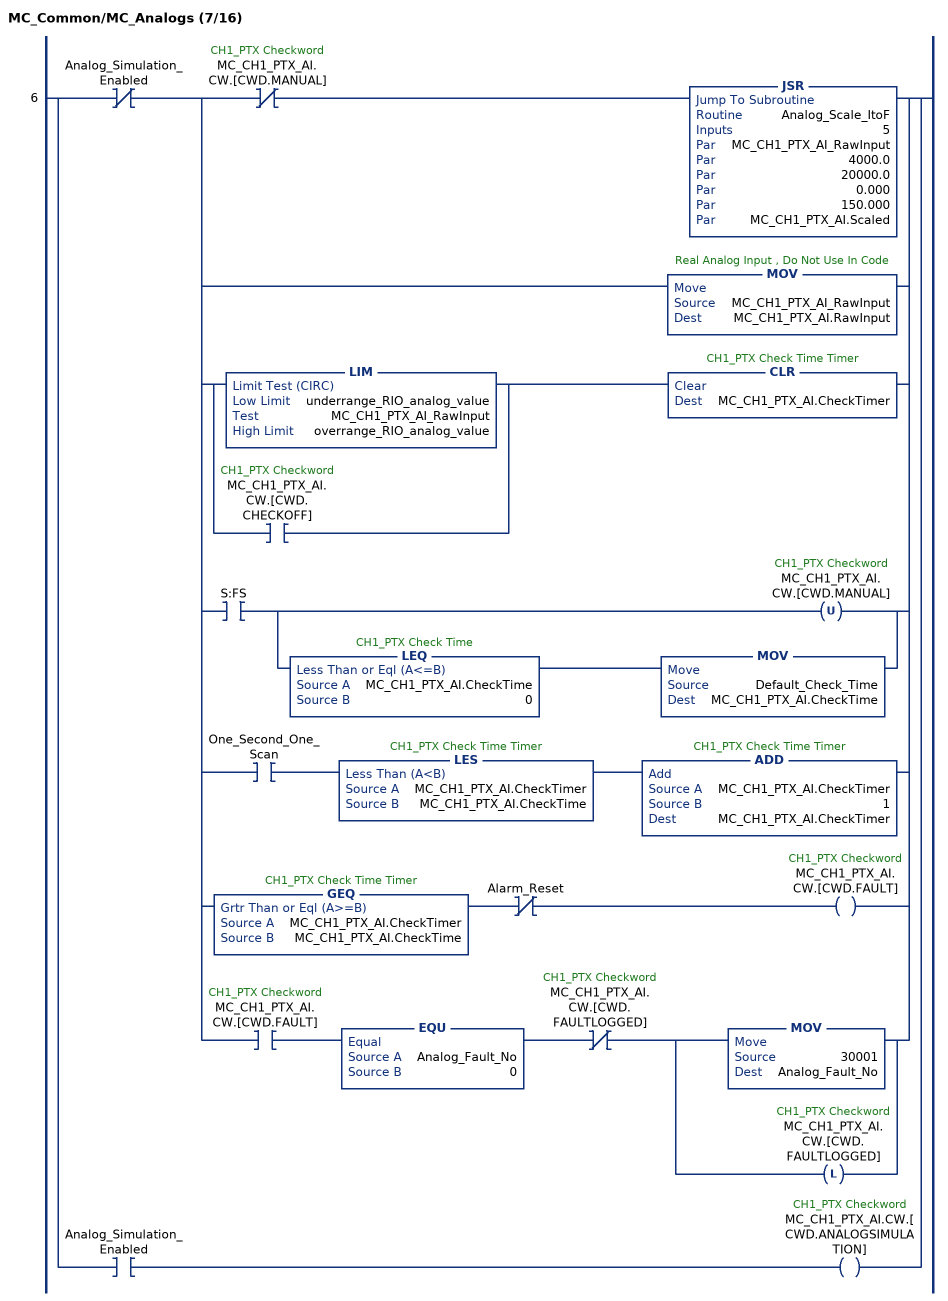
   6: [XIO(Analog_Simulation_Enabled) [XIO(MC_CH1_PTX_AI.CW.[CWD.MANUAL]) JSR(Analog_Scale_ItoF,5,MC_CH1_PTX_AI_RawInput,4000.0,20000.0,0.000,150.000,MC_CH1_PTX_AI.Scaled) ,MOV(MC_CH1_PTX_AI_RawInput,MC_CH1_PTX_AI.RawInput) ,[LIM(underrange_RIO_analog_value,MC_CH1_PTX_AI_RawInput,overrange_RIO_analog_value) ,XIC(MC_CH1_PTX_AI.CW.[CWD.CHECKOFF]) ] CLR(MC_CH1_PTX_AI.CheckTimer) ,XIC(S:FS) [OTU(MC_CH1_PTX_AI.CW.[CWD.MANUAL]) ,LEQ(MC_CH1_PTX_AI.CheckTime,0) MOV(Default_Check_Time,MC_CH1_PTX_AI.CheckTime) ] ,XIC(One_Second_One_Scan) LES(MC_CH1_PTX_AI.CheckTimer,MC_CH1_PTX_AI.CheckTime) ADD(MC_CH1_PTX_AI.CheckTimer,1,MC_CH1_PTX_AI.CheckTimer) ,GEQ(MC_CH1_PTX_AI.CheckTimer,MC_CH1_PTX_AI.CheckTime) XIO(Alarm_Reset) OTE(MC_CH1_PTX_AI.CW.[CWD.FAULT]) ,XIC(MC_CH1_PTX_AI.CW.[CWD.FAULT]) EQU(Analog_Fault_No,0) XIO(MC_CH1_PTX_AI.CW.[CWD.FAULTLOGGED]) [MOV(30001,Analog_Fault_No) ,OTL(MC_CH1_PTX_AI.CW.[CWD.FAULTLOGGED]) ] ] ,XIC(Analog_Simulation_Enabled) OTE(MC_CH1_PTX_AI.CW.[CWD.ANALOGSIMULATION]) ];
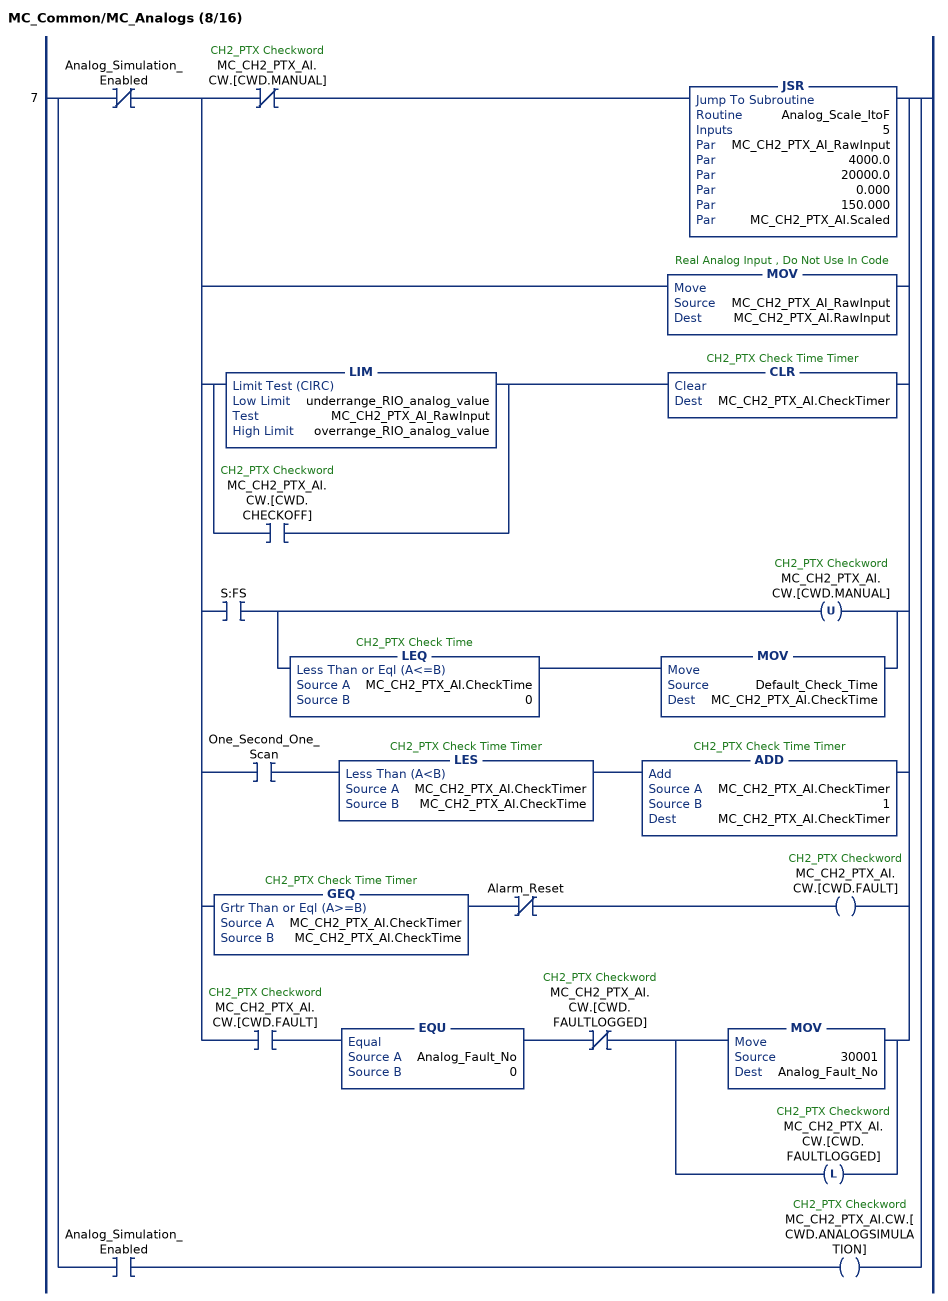
   7: [XIO(Analog_Simulation_Enabled) [XIO(MC_CH2_PTX_AI.CW.[CWD.MANUAL]) JSR(Analog_Scale_ItoF,5,MC_CH2_PTX_AI_RawInput,4000.0,20000.0,0.000,150.000,MC_CH2_PTX_AI.Scaled) ,MOV(MC_CH2_PTX_AI_RawInput,MC_CH2_PTX_AI.RawInput) ,[LIM(underrange_RIO_analog_value,MC_CH2_PTX_AI_RawInput,overrange_RIO_analog_value) ,XIC(MC_CH2_PTX_AI.CW.[CWD.CHECKOFF]) ] CLR(MC_CH2_PTX_AI.CheckTimer) ,XIC(S:FS) [OTU(MC_CH2_PTX_AI.CW.[CWD.MANUAL]) ,LEQ(MC_CH2_PTX_AI.CheckTime,0) MOV(Default_Check_Time,MC_CH2_PTX_AI.CheckTime) ] ,XIC(One_Second_One_Scan) LES(MC_CH2_PTX_AI.CheckTimer,MC_CH2_PTX_AI.CheckTime) ADD(MC_CH2_PTX_AI.CheckTimer,1,MC_CH2_PTX_AI.CheckTimer) ,GEQ(MC_CH2_PTX_AI.CheckTimer,MC_CH2_PTX_AI.CheckTime) XIO(Alarm_Reset) OTE(MC_CH2_PTX_AI.CW.[CWD.FAULT]) ,XIC(MC_CH2_PTX_AI.CW.[CWD.FAULT]) EQU(Analog_Fault_No,0) XIO(MC_CH2_PTX_AI.CW.[CWD.FAULTLOGGED]) [MOV(30001,Analog_Fault_No) ,OTL(MC_CH2_PTX_AI.CW.[CWD.FAULTLOGGED]) ] ] ,XIC(Analog_Simulation_Enabled) OTE(MC_CH2_PTX_AI.CW.[CWD.ANALOGSIMULATION]) ];
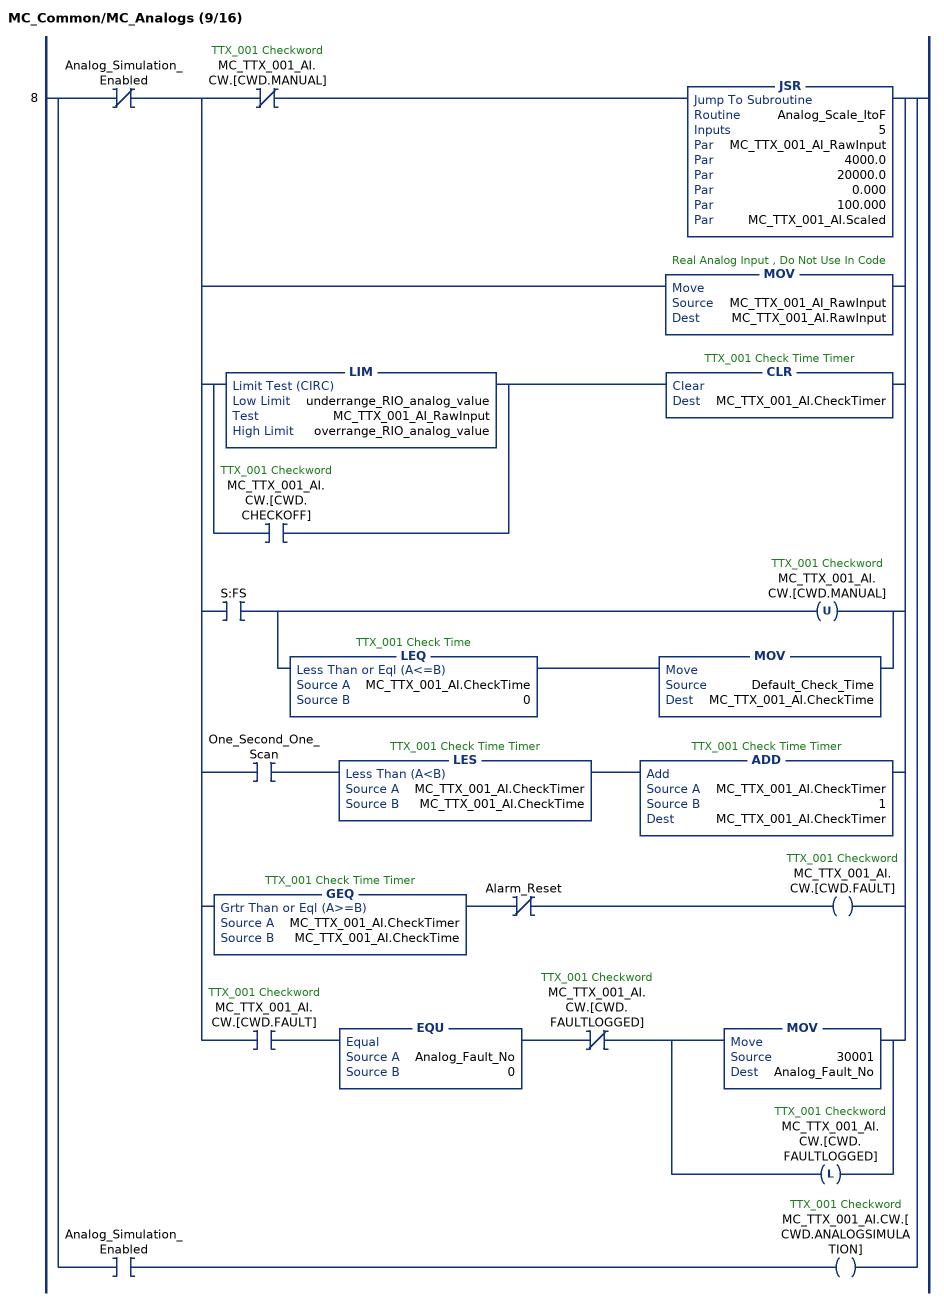
   8: [XIO(Analog_Simulation_Enabled) [XIO(MC_TTX_001_AI.CW.[CWD.MANUAL]) JSR(Analog_Scale_ItoF,5,MC_TTX_001_AI_RawInput,4000.0,20000.0,0.000,100.000,MC_TTX_001_AI.Scaled) ,MOV(MC_TTX_001_AI_RawInput,MC_TTX_001_AI.RawInput) ,[LIM(underrange_RIO_analog_value,MC_TTX_001_AI_RawInput,overrange_RIO_analog_value) ,XIC(MC_TTX_001_AI.CW.[CWD.CHECKOFF]) ] CLR(MC_TTX_001_AI.CheckTimer) ,XIC(S:FS) [OTU(MC_TTX_001_AI.CW.[CWD.MANUAL]) ,LEQ(MC_TTX_001_AI.CheckTime,0) MOV(Default_Check_Time,MC_TTX_001_AI.CheckTime) ] ,XIC(One_Second_One_Scan) LES(MC_TTX_001_AI.CheckTimer,MC_TTX_001_AI.CheckTime) ADD(MC_TTX_001_AI.CheckTimer,1,MC_TTX_001_AI.CheckTimer) ,GEQ(MC_TTX_001_AI.CheckTimer,MC_TTX_001_AI.CheckTime) XIO(Alarm_Reset) OTE(MC_TTX_001_AI.CW.[CWD.FAULT]) ,XIC(MC_TTX_001_AI.CW.[CWD.FAULT]) EQU(Analog_Fault_No,0) XIO(MC_TTX_001_AI.CW.[CWD.FAULTLOGGED]) [MOV(30001,Analog_Fault_No) ,OTL(MC_TTX_001_AI.CW.[CWD.FAULTLOGGED]) ] ] ,XIC(Analog_Simulation_Enabled) OTE(MC_TTX_001_AI.CW.[CWD.ANALOGSIMULATION]) ];
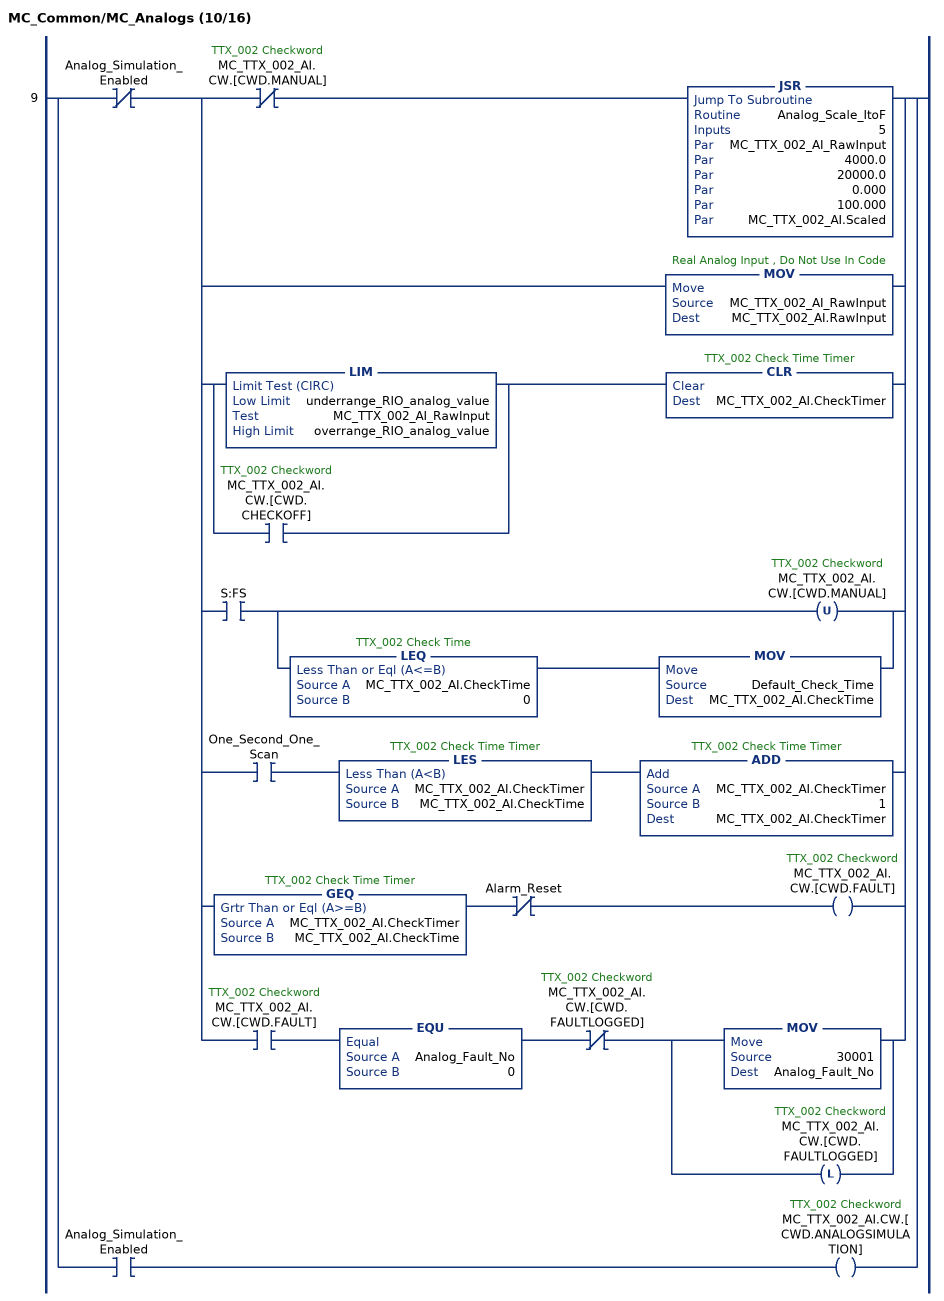
   9: [XIO(Analog_Simulation_Enabled) [XIO(MC_TTX_002_AI.CW.[CWD.MANUAL]) JSR(Analog_Scale_ItoF,5,MC_TTX_002_AI_RawInput,4000.0,20000.0,0.000,100.000,MC_TTX_002_AI.Scaled) ,MOV(MC_TTX_002_AI_RawInput,MC_TTX_002_AI.RawInput) ,[LIM(underrange_RIO_analog_value,MC_TTX_002_AI_RawInput,overrange_RIO_analog_value) ,XIC(MC_TTX_002_AI.CW.[CWD.CHECKOFF]) ] CLR(MC_TTX_002_AI.CheckTimer) ,XIC(S:FS) [OTU(MC_TTX_002_AI.CW.[CWD.MANUAL]) ,LEQ(MC_TTX_002_AI.CheckTime,0) MOV(Default_Check_Time,MC_TTX_002_AI.CheckTime) ] ,XIC(One_Second_One_Scan) LES(MC_TTX_002_AI.CheckTimer,MC_TTX_002_AI.CheckTime) ADD(MC_TTX_002_AI.CheckTimer,1,MC_TTX_002_AI.CheckTimer) ,GEQ(MC_TTX_002_AI.CheckTimer,MC_TTX_002_AI.CheckTime) XIO(Alarm_Reset) OTE(MC_TTX_002_AI.CW.[CWD.FAULT]) ,XIC(MC_TTX_002_AI.CW.[CWD.FAULT]) EQU(Analog_Fault_No,0) XIO(MC_TTX_002_AI.CW.[CWD.FAULTLOGGED]) [MOV(30001,Analog_Fault_No) ,OTL(MC_TTX_002_AI.CW.[CWD.FAULTLOGGED]) ] ] ,XIC(Analog_Simulation_Enabled) OTE(MC_TTX_002_AI.CW.[CWD.ANALOGSIMULATION]) ];
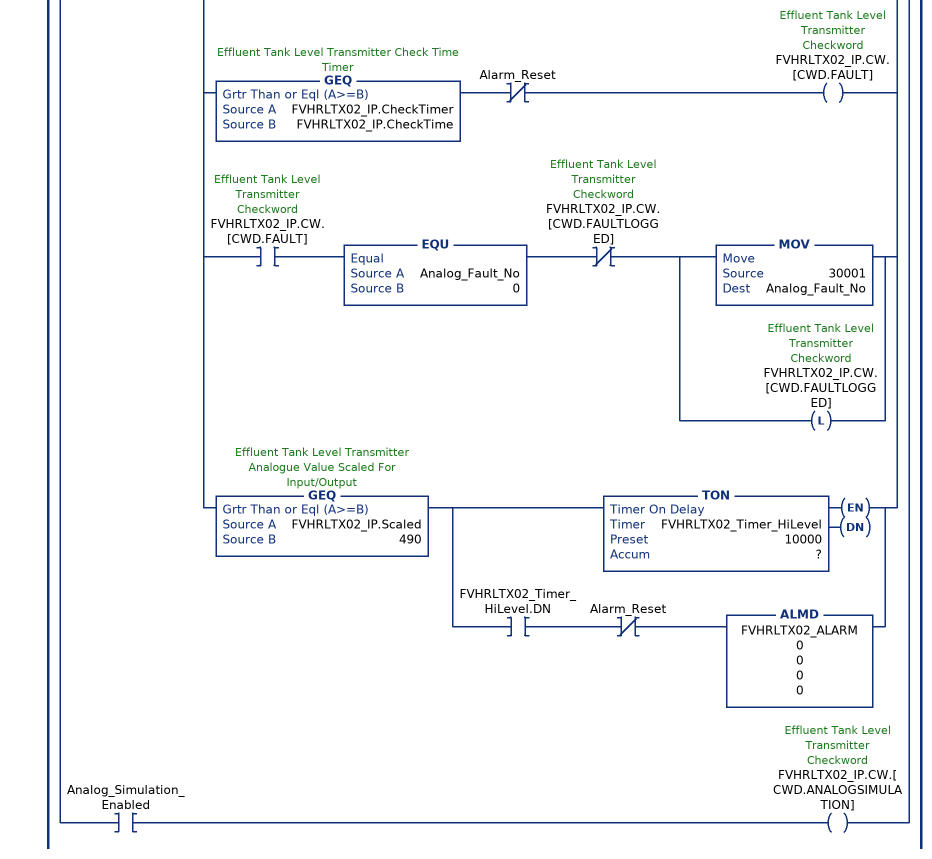
   10: [XIO(Analog_Simulation_Enabled) [XIO(FVHRLTX02_IP.CW.[CWD.MANUAL]) [JSR(Analog_Scale_ItoF,5,FVHRLTX02_IP_RawInput,4000.0,20000.0,0.0,500.0,FVHRLTX02_IP.Scaled) ,CPT(FVHRLTX02_IP_Percentage,(FVHRLTX02_IP.Scaled / 500) * 100) ] ,MOV(FVHRLTX02_IP_RawInput,FVHRLTX02_IP.RawInput) ,[LIM(underrange_RIO_analog_value,FVHRLTX02_IP_RawInput,overrange_RIO_analog_value) ,XIC(FVHRLTX02_IP.CW.[CWD.CHECKOFF]) ] CLR(FVHRLTX02_IP.CheckTimer) ,XIC(S:FS) [OTU(FVHRLTX02_IP.CW.[CWD.MANUAL]) ,LEQ(FVHRLTX02_IP.CheckTime,0) MOV(Default_Check_Time,FVHRLTX02_IP.CheckTime) ] ,XIC(One_Second_One_Scan) LES(FVHRLTX02_IP.CheckTimer,FVHRLTX02_IP.CheckTime) ADD(FVHRLTX02_IP.CheckTimer,1,FVHRLTX02_IP.CheckTimer) ,GEQ(FVHRLTX02_IP.CheckTimer,FVHRLTX02_IP.CheckTime) XIO(Alarm_Reset) OTE(FVHRLTX02_IP.CW.[CWD.FAULT]) ,XIC(FVHRLTX02_IP.CW.[CWD.FAULT]) EQU(Analog_Fault_No,0) XIO(FVHRLTX02_IP.CW.[CWD.FAULTLOGGED]) [MOV(30001,Analog_Fault_No) ,OTL(FVHRLTX02_IP.CW.[CWD.FAULTLOGGED]) ] ,GEQ(FVHRLTX02_IP.Scaled,490) [TON(FVHRLTX02_Timer_HiLevel,?,?) ,XIC(FVHRLTX02_Timer_HiLevel.DN) XIO(Alarm_Reset) ALMD(FVHRLTX02_ALARM,0,0,0,0) ] ] ,XIC(Analog_Simulation_Enabled) OTE(FVHRLTX02_IP.CW.[CWD.ANALOGSIMULATION]) ];
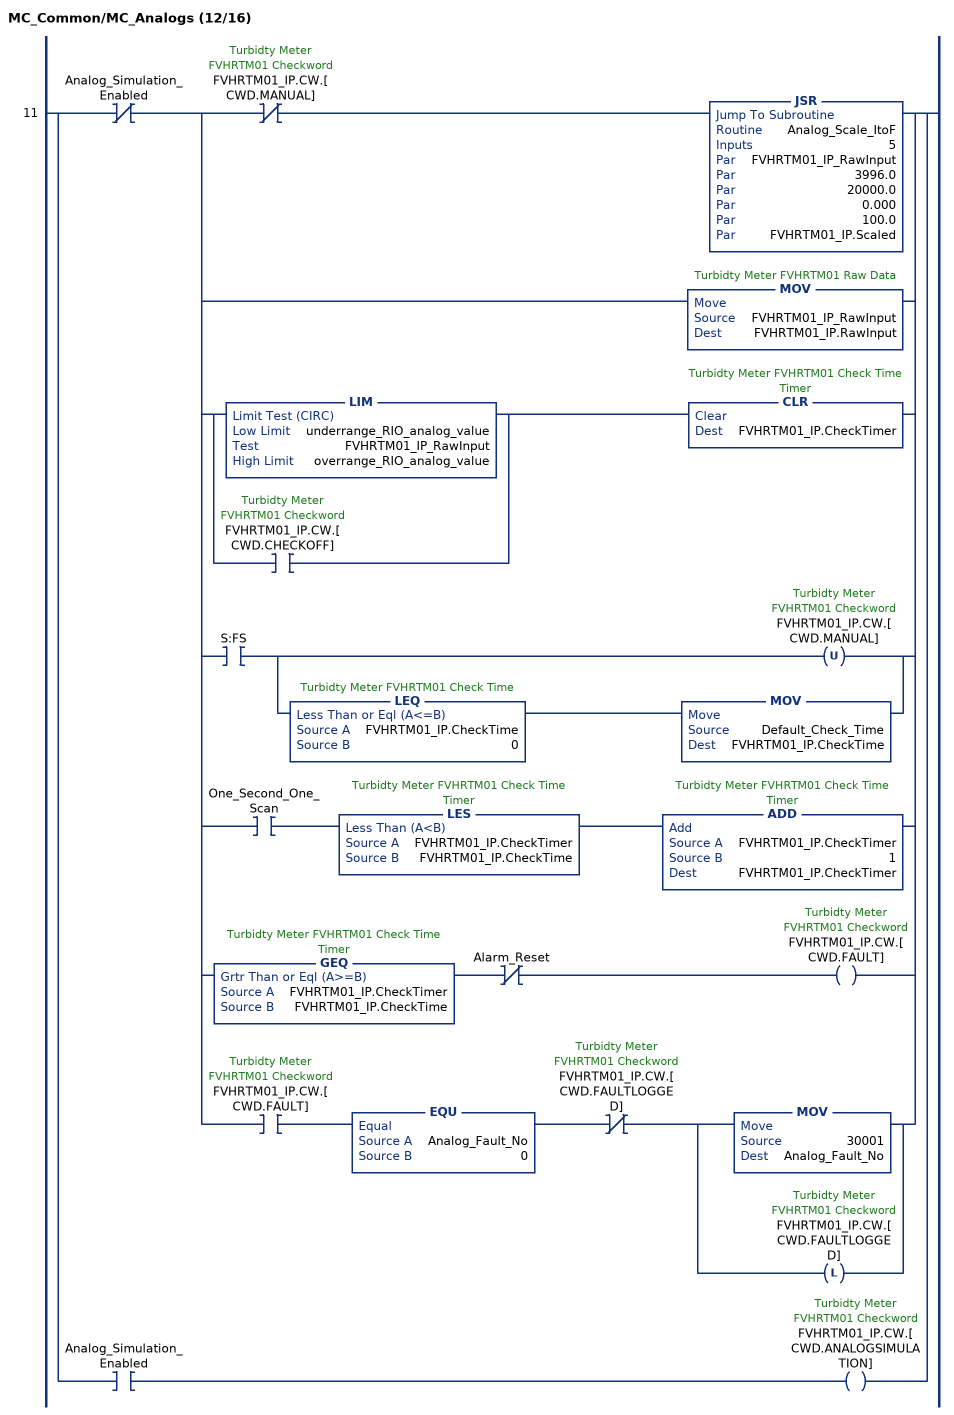
   11: [XIO(Analog_Simulation_Enabled) [XIO(FVHRTM01_IP.CW.[CWD.MANUAL]) JSR(Analog_Scale_ItoF,5,FVHRTM01_IP_RawInput,3996.0,20000.0,0.000,100.0,FVHRTM01_IP.Scaled) ,MOV(FVHRTM01_IP_RawInput,FVHRTM01_IP.RawInput) ,[LIM(underrange_RIO_analog_value,FVHRTM01_IP_RawInput,overrange_RIO_analog_value) ,XIC(FVHRTM01_IP.CW.[CWD.CHECKOFF]) ] CLR(FVHRTM01_IP.CheckTimer) ,XIC(S:FS) [OTU(FVHRTM01_IP.CW.[CWD.MANUAL]) ,LEQ(FVHRTM01_IP.CheckTime,0) MOV(Default_Check_Time,FVHRTM01_IP.CheckTime) ] ,XIC(One_Second_One_Scan) LES(FVHRTM01_IP.CheckTimer,FVHRTM01_IP.CheckTime) ADD(FVHRTM01_IP.CheckTimer,1,FVHRTM01_IP.CheckTimer) ,GEQ(FVHRTM01_IP.CheckTimer,FVHRTM01_IP.CheckTime) XIO(Alarm_Reset) OTE(FVHRTM01_IP.CW.[CWD.FAULT]) ,XIC(FVHRTM01_IP.CW.[CWD.FAULT]) EQU(Analog_Fault_No,0) XIO(FVHRTM01_IP.CW.[CWD.FAULTLOGGED]) [MOV(30001,Analog_Fault_No) ,OTL(FVHRTM01_IP.CW.[CWD.FAULTLOGGED]) ] ] ,XIC(Analog_Simulation_Enabled) OTE(FVHRTM01_IP.CW.[CWD.ANALOGSIMULATION]) ];
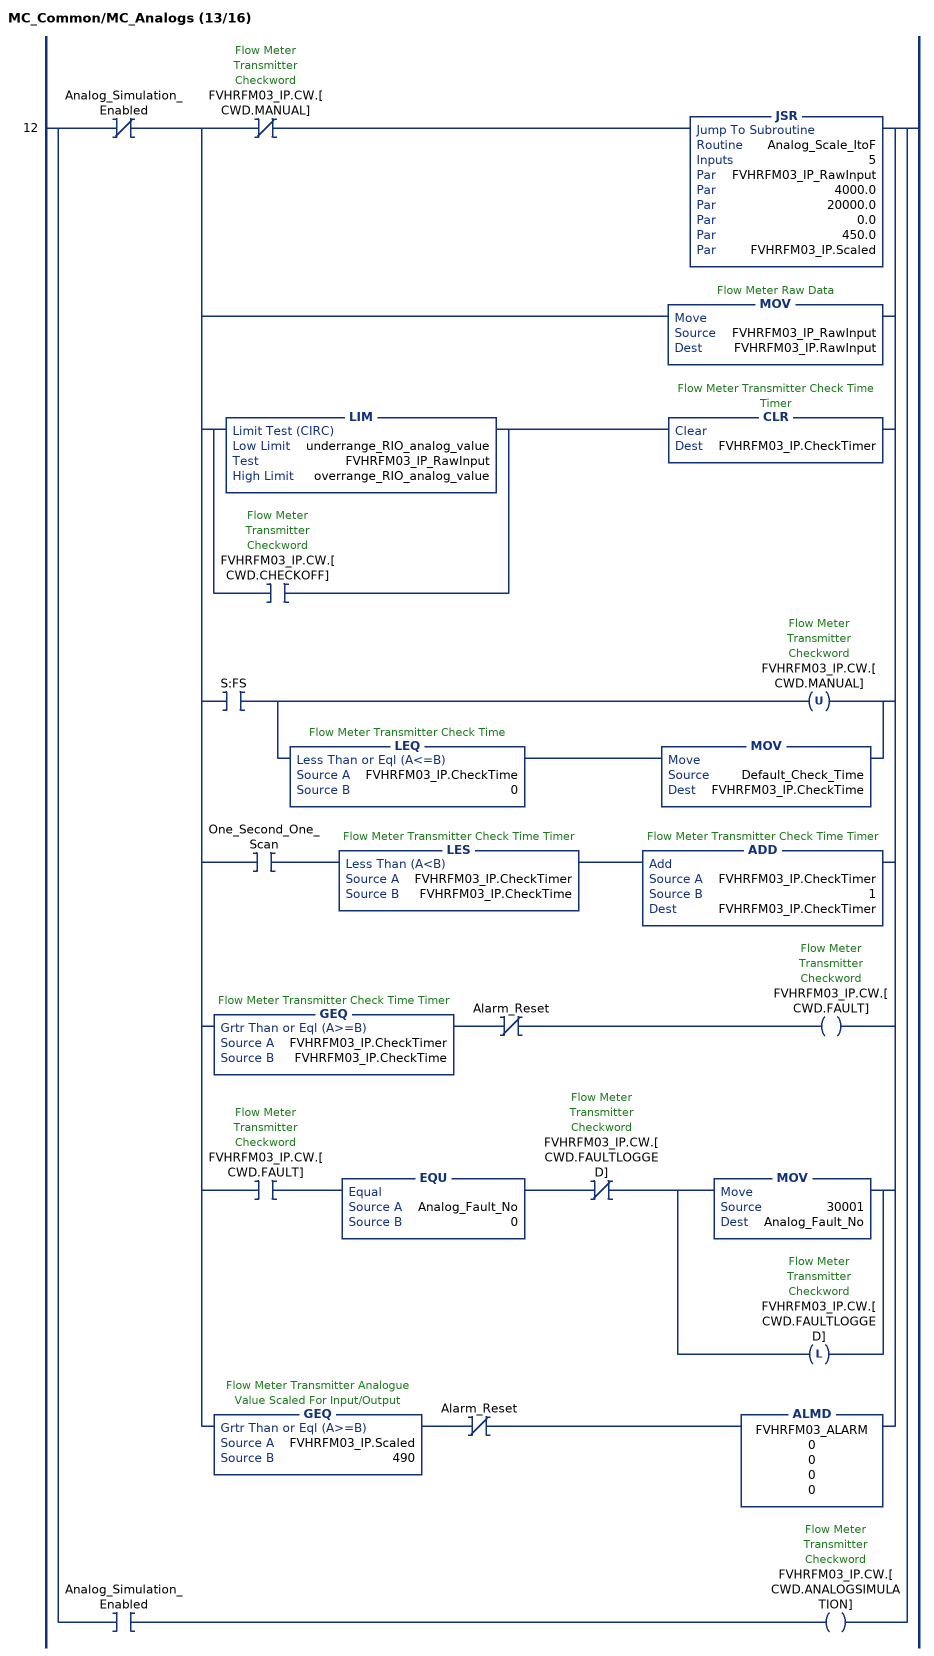
   12: [XIO(Analog_Simulation_Enabled) [XIO(FVHRFM03_IP.CW.[CWD.MANUAL]) JSR(Analog_Scale_ItoF,5,FVHRFM03_IP_RawInput,4000.0,20000.0,0.0,450.0,FVHRFM03_IP.Scaled) ,MOV(FVHRFM03_IP_RawInput,FVHRFM03_IP.RawInput) ,[LIM(underrange_RIO_analog_value,FVHRFM03_IP_RawInput,overrange_RIO_analog_value) ,XIC(FVHRFM03_IP.CW.[CWD.CHECKOFF]) ] CLR(FVHRFM03_IP.CheckTimer) ,XIC(S:FS) [OTU(FVHRFM03_IP.CW.[CWD.MANUAL]) ,LEQ(FVHRFM03_IP.CheckTime,0) MOV(Default_Check_Time,FVHRFM03_IP.CheckTime) ] ,XIC(One_Second_One_Scan) LES(FVHRFM03_IP.CheckTimer,FVHRFM03_IP.CheckTime) ADD(FVHRFM03_IP.CheckTimer,1,FVHRFM03_IP.CheckTimer) ,GEQ(FVHRFM03_IP.CheckTimer,FVHRFM03_IP.CheckTime) XIO(Alarm_Reset) OTE(FVHRFM03_IP.CW.[CWD.FAULT]) ,XIC(FVHRFM03_IP.CW.[CWD.FAULT]) EQU(Analog_Fault_No,0) XIO(FVHRFM03_IP.CW.[CWD.FAULTLOGGED]) [MOV(30001,Analog_Fault_No) ,OTL(FVHRFM03_IP.CW.[CWD.FAULTLOGGED]) ] ,GEQ(FVHRFM03_IP.Scaled,490) XIO(Alarm_Reset) ALMD(FVHRFM03_ALARM,0,0,0,0) ] ,XIC(Analog_Simulation_Enabled) OTE(FVHRFM03_IP.CW.[CWD.ANALOGSIMULATION]) ];
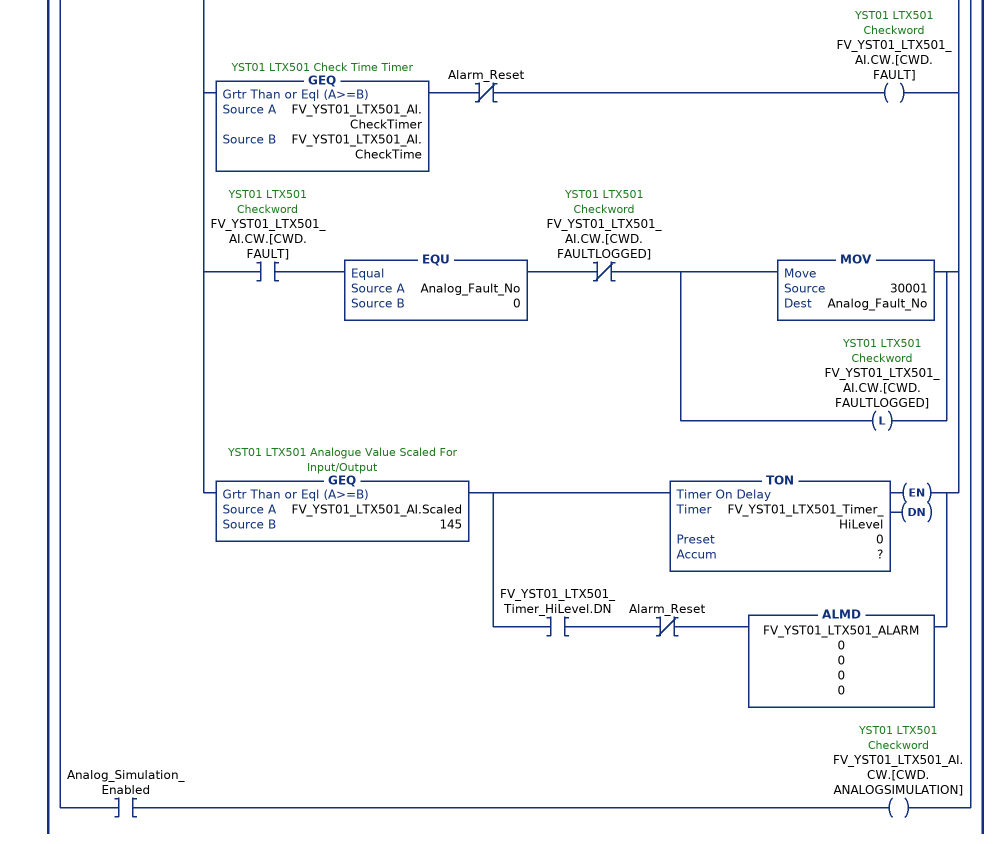
   13: [XIO(Analog_Simulation_Enabled) [XIO(FV_YST01_LTX501_AI.CW.[CWD.MANUAL]) JSR(Analog_Scale_ItoF,5,FV_YST01_LTX501_AI_RawInput,4000.0,20000.0,0.0,150.0,FV_YST01_LTX501_AI.Scaled) ,MOV(FV_YST01_LTX501_AI.Scaled,YST_Data[0]) ,MOV(FV_YST01_LTX501_AI_RawInput,FV_YST01_LTX501_AI.RawInput) ,[LIM(underrange_RIO_analog_value,FV_YST01_LTX501_AI_RawInput,overrange_RIO_analog_value) ,XIC(FV_YST01_LTX501_AI.CW.[CWD.CHECKOFF]) ] CLR(FV_YST01_LTX501_AI.CheckTimer) ,XIC(S:FS) [OTU(FV_YST01_LTX501_AI.CW.[CWD.MANUAL]) ,LEQ(FV_YST01_LTX501_AI.CheckTime,0) MOV(Default_Check_Time,FV_YST01_LTX501_AI.CheckTime) ] ,XIC(One_Second_One_Scan) LES(FV_YST01_LTX501_AI.CheckTimer,FV_YST01_LTX501_AI.CheckTime) ADD(FV_YST01_LTX501_AI.CheckTimer,1,FV_YST01_LTX501_AI.CheckTimer) ,GEQ(FV_YST01_LTX501_AI.CheckTimer,FV_YST01_LTX501_AI.CheckTime) XIO(Alarm_Reset) OTE(FV_YST01_LTX501_AI.CW.[CWD.FAULT]) ,XIC(FV_YST01_LTX501_AI.CW.[CWD.FAULT]) EQU(Analog_Fault_No,0) XIO(FV_YST01_LTX501_AI.CW.[CWD.FAULTLOGGED]) [MOV(30001,Analog_Fault_No) ,OTL(FV_YST01_LTX501_AI.CW.[CWD.FAULTLOGGED]) ] ,GEQ(FV_YST01_LTX501_AI.Scaled,145) [TON(FV_YST01_LTX501_Timer_HiLevel,?,?) ,XIC(FV_YST01_LTX501_Timer_HiLevel.DN) XIO(Alarm_Reset) ALMD(FV_YST01_LTX501_ALARM,0,0,0,0) ] ] ,XIC(Analog_Simulation_Enabled) OTE(FV_YST01_LTX501_AI.CW.[CWD.ANALOGSIMULATION]) ];
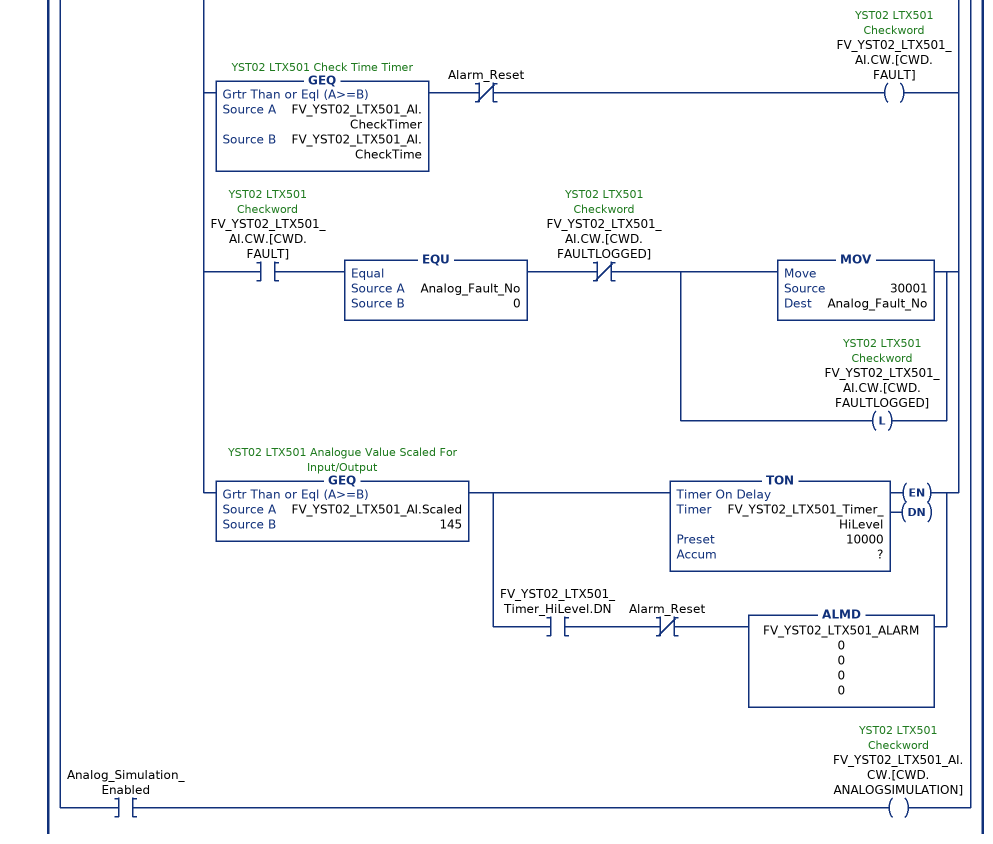
   14: [XIO(Analog_Simulation_Enabled) [XIO(FV_YST02_LTX501_AI.CW.[CWD.MANUAL]) JSR(Analog_Scale_ItoF,5,FV_YST02_LTX501_AI_RawInput,4000.0,20000.0,0.0,150.0,FV_YST02_LTX501_AI.Scaled) ,MOV(FV_YST02_LTX501_AI.Scaled,YST_Data[1]) ,MOV(FV_YST02_LTX501_AI_RawInput,FV_YST02_LTX501_AI.RawInput) ,[LIM(underrange_RIO_analog_value,FV_YST02_LTX501_AI_RawInput,overrange_RIO_analog_value) ,XIC(FV_YST02_LTX501_AI.CW.[CWD.CHECKOFF]) ] CLR(FV_YST02_LTX501_AI.CheckTimer) ,XIC(S:FS) [OTU(FV_YST02_LTX501_AI.CW.[CWD.MANUAL]) ,LEQ(FV_YST02_LTX501_AI.CheckTime,0) MOV(Default_Check_Time,FV_YST02_LTX501_AI.CheckTime) ] ,XIC(One_Second_One_Scan) LES(FV_YST02_LTX501_AI.CheckTimer,FV_YST02_LTX501_AI.CheckTime) ADD(FV_YST02_LTX501_AI.CheckTimer,1,FV_YST02_LTX501_AI.CheckTimer) ,GEQ(FV_YST02_LTX501_AI.CheckTimer,FV_YST02_LTX501_AI.CheckTime) XIO(Alarm_Reset) OTE(FV_YST02_LTX501_AI.CW.[CWD.FAULT]) ,XIC(FV_YST02_LTX501_AI.CW.[CWD.FAULT]) EQU(Analog_Fault_No,0) XIO(FV_YST02_LTX501_AI.CW.[CWD.FAULTLOGGED]) [MOV(30001,Analog_Fault_No) ,OTL(FV_YST02_LTX501_AI.CW.[CWD.FAULTLOGGED]) ] ,GEQ(FV_YST02_LTX501_AI.Scaled,145) [TON(FV_YST02_LTX501_Timer_HiLevel,?,?) ,XIC(FV_YST02_LTX501_Timer_HiLevel.DN) XIO(Alarm_Reset) ALMD(FV_YST02_LTX501_ALARM,0,0,0,0) ] ] ,XIC(Analog_Simulation_Enabled) OTE(FV_YST02_LTX501_AI.CW.[CWD.ANALOGSIMULATION]) ];
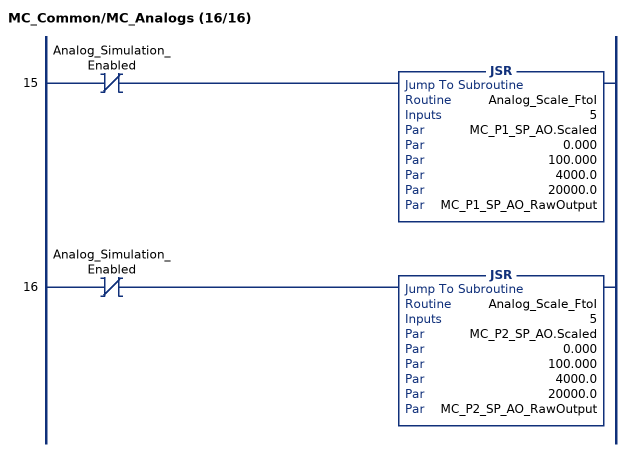
   15: XIO(Analog_Simulation_Enabled)JSR(Analog_Scale_FtoI,5,MC_P1_SP_AO.Scaled,0.000,100.000,4000.0,20000.0,MC_P1_SP_AO_RawOutput);
   16: XIO(Analog_Simulation_Enabled)JSR(Analog_Scale_FtoI,5,MC_P2_SP_AO.Scaled,0.000,100.000,4000.0,20000.0,MC_P2_SP_AO_RawOutput);
END_ROUTINE
